// TIA Portal project "maupTIA_DEMO2023_V17" (V17) (continued)

       END_IF;
       #DrainingPhase.Cmd.StartMan := FALSE;
       #DrainingPhase.Cmd.PauseMan := FALSE;
       #DrainingPhase.Cmd.ResumeMan := FALSE;
       #DrainingPhase.Cmd.StopMan := FALSE;
   END_REGION

   REGION AutCtrl
       //if request to run in automatic mode -> set auto request to open of filling valve to 1 and close to 0, if not open 0 close 1
       // commands should be sets to false after their processing
       IF #DrainingPhase.State.AutCtrl THEN
           IF #DrainingPhase.Cmd.StartAut THEN
               #DrainingPhase.State.Running := TRUE;
               #DrainingPhase.State.Idle := FALSE;

               #DrainingPhase.Cmd.StartAut := FALSE;

               #DrainingValve.Cmd.AutCtrl := TRUE;




           END_IF;

           IF #DrainingPhase.Cmd.StopAut THEN
               #DrainingPhase.State.Running := FALSE;
               #DrainingPhase.State.Idle := TRUE;

               #DrainingPhase.Cmd.StopAut := FALSE;


           END_IF;

       END_IF;
   END_REGION

   REGION Done
       //every phase should have finish condition - draining phase - if water level is below requested level
       //after that done state should be setted to 1
       #DrainingPhase.Param.DrainLevel := 0.01;
       IF #DrainingPhase.WaterLevel <= #DrainingPhase.Param.DrainLevel THEN // kdyz je vypusteno, mozna je to zase ta promenna ktere preteka, nvm
           #DrainingPhase.Cmd.StopAut := TRUE;
           #DrainingPhase.Cmd.StopMan := TRUE;
           #DrainingPhase.State.Done := TRUE;
       END_IF;

       // command reset done resets done state and than resets command

       IF #DrainingPhase.Cmd.ResetDone THEN // AND DONE = TRUE? mozna zbytecne.
           #DrainingPhase.State.Done := FALSE;
           #DrainingPhase.Cmd.ResetDone := FALSE;
       END_IF;

   END_REGION

   REGION States 
       //Command valve in cases of states
       IF #DrainingPhase.State.Running THEN
           #DrainingValve.Cmd.Req2OpenAut := TRUE;
           #DrainingValve.Cmd.Req2CloseAut := FALSE;
          // #DrainingValve.Cmd.Req2CloseAut := FALSE;
       ELSE
           #DrainingValve.Cmd.Req2OpenAut := FALSE;
           #DrainingValve.Cmd.Req2CloseAut := TRUE;
           //#DrainingValve.Cmd.Req2CloseAut := FALSE;
       END_IF;
   END_REGION

   // delault state of phase - if not any state sets state to idle
   IF NOT #DrainingPhase.State.Idle AND NOT #DrainingPhase.State.Paused AND NOT #DrainingPhase.State.Running THEN
       #DrainingPhase.State.Idle := TRUE;
   END_IF;

   IF #DrainingPhase.State.Running THEN
       #DrainingPhase.State.StateInt := #Running;
   ELSIF #DrainingPhase.State.Paused THEN
       #DrainingPhase.State.StateInt := #Pause;
   ELSIF #DrainingPhase.State.Idle THEN
       #DrainingPhase.State.StateInt := #Idle;
   ELSIF #DrainingPhase.State.Done THEN
       #DrainingPhase.State.StateInt := #Idle;
   END_IF;
END_FUNCTION_BLOCK

FUNCTION_BLOCK "MixingFC"   // FB6, SCL
{ S7_Optimized_Access := 'TRUE' }
VERSION : 0.1
   VAR_IN_OUT
      MixingPhase : "PhaseMixing";
      MixerEng : "Engine";
   END_VAR
   VAR
      fElapsedTime : Int;
      fSecImp : R_TRIG;
   END_VAR
   VAR_TEMP
      tmp : Bool;
   END_VAR
   VAR CONSTANT
      Idle : Int := 0;
      Running : Int := 1;
      Pause : Int := 2;
   END_VAR
BEGIN
   REGION Aut/Man
       // switching state of engine - automatic or manual control (default state is manual)
       IF #MixingPhase.Cmd.AutCtrl THEN
           #MixingPhase.State.ManCtrl := FALSE;
           #MixingPhase.State.AutCtrl := TRUE;
           #MixingPhase.Cmd.AutCtrl := FALSE;
       END_IF;

       IF #MixingPhase.Cmd.ManCtrl THEN
           #MixingPhase.State.AutCtrl := FALSE;
           #MixingPhase.State.ManCtrl := TRUE;
           #MixingPhase.Cmd.ManCtrl := FALSE;
       END_IF;

       IF NOT #MixingPhase.State.AutCtrl AND NOT #MixingPhase.State.ManCtrl THEN
           #MixingPhase.State.ManCtrl := TRUE; // nebo dat Cmd.Manctrl do TRUE aby prosel IF nahore?
       END_IF;

   END_REGION

   REGION ManCtrl
       // processing manual actions - if command is processed, it is sets to FALSE even if can't be processed
       // Phase commands are start, stop, pause and resume 
       // Start - start mixing  
       // Stop - stop mixing
       // Pause - stop mixing 
       // Resume - start mixing
       // real states of phase are writed into states in phase structure

       IF #MixingPhase.State.ManCtrl THEN
           IF #MixingPhase.Cmd.StartMan THEN
               #MixingPhase.State.Paused := FALSE;
               #MixingPhase.State.Idle := FALSE;
               #MixingPhase.State.Running := TRUE;

               #MixerEng.Cmd.TurnOnMan := TRUE;
               //#MixerEng.Cmd.TurnOnMan := FALSE;

               #MixingPhase.Cmd.ResetDone := TRUE;
               //#MixingPhase.Cmd.ResetDone := FALSE;
           END_IF;

           IF #MixingPhase.State.Running THEN
               IF #MixingPhase.Cmd.PauseMan THEN
                   #MixingPhase.State.Running := FALSE;
                   #MixingPhase.State.Idle := FALSE;
                   #MixingPhase.State.Paused := TRUE;

                   #MixerEng.Cmd.TurnOffMan := TRUE;
                  // #MixerEng.Cmd.TurnOffMan := FALSE;

                   #MixingPhase.Cmd.ResetDone := TRUE;
                   //#MixingPhase.Cmd.ResetDone := FALSE;
               END_IF;
           END_IF;

           IF #MixingPhase.State.Paused THEN
               IF #MixingPhase.Cmd.ResumeMan THEN
                   #MixingPhase.State.Paused := FALSE;
                   #MixingPhase.State.Idle := FALSE;
                   #MixingPhase.State.Running := TRUE;

                   #MixerEng.Cmd.TurnOnMan := TRUE;
                   //#MixerEng.Cmd.TurnOnMan := FALSE;

                   #MixingPhase.Cmd.ResetDone := TRUE;
                   //#MixingPhase.Cmd.ResetDone := FALSE;
               END_IF;
           END_IF;


           IF #MixingPhase.State.Running OR #MixingPhase.State.Paused THEN
               IF #MixingPhase.Cmd.StopMan THEN
                   #MixingPhase.State.Running := FALSE;
                   #MixingPhase.State.Paused := FALSE;
                   #MixingPhase.State.Idle := TRUE;

                   #MixerEng.Cmd.TurnOffMan := TRUE;
                   //#MixerEng.Cmd.TurnOffMan := FALSE;

                   #MixingPhase.Cmd.ResetDone := TRUE;
                   //#MixingPhase.Cmd.ResetDone := FALSE;
               END_IF;
           END_IF;


       END_IF;
       #MixingPhase.Cmd.StartMan := FALSE;
       #MixingPhase.Cmd.PauseMan := FALSE;
       #MixingPhase.Cmd.ResumeMan := FALSE;
       #MixingPhase.Cmd.StopMan := FALSE;
   END_REGION

   REGION AutCtrl
       // if request to run in automatic mode -> set auto request to mixing to 1, if not request to mixing is 0
       // commands should be sets to false after their processing
       IF #MixingPhase.State.AutCtrl THEN
           IF #MixingPhase.Cmd.StartAut THEN
               #MixingPhase.State.Running := TRUE;
               #MixingPhase.State.Idle := FALSE;
               #MixingPhase.Cmd.StartAut := FALSE;
               #MixerEng.Cmd.AutCtrl := TRUE;
           END_IF;

           IF #MixingPhase.Cmd.StopAut THEN
               #MixingPhase.State.Running := FALSE;
               #MixingPhase.State.Idle := TRUE;
               #MixingPhase.Cmd.StopAut := FALSE;
           END_IF;

       END_IF;

   END_REGION


   REGION Done
       // every phase should have finish condition - mixing phase - if time of runnig is bigger or same as requested
       // after that done state should be setted to 1

       // command reset done resets done state and than resets command
       // calculation of elapsed time from engin state RT
       IF #MixingPhase.State.Running THEN
           "fSecImp"(CLK := "Clock_1Hz",
                     Q => #tmp);
           IF #tmp THEN
               #fElapsedTime := #fElapsedTime + 1;
           END_IF;

       END_IF;

       IF #MixingPhase.Param.TimeSec <= #fElapsedTime THEN // kdyz je domixovano, mozna je to zase ta promenna ktere preteka, nvm
           #MixingPhase.Cmd.StopAut := TRUE;
           #MixingPhase.Cmd.StopMan := TRUE;
           #MixingPhase.State.Done := TRUE;
       END_IF;


       // command reset done resets done state and than resets command
       IF #MixingPhase.Cmd.ResetDone THEN // AND DONE = TRUE? mozna zbytecne.
           // reset timer
           #MixingPhase.State.Done := FALSE;
           #fElapsedTime := 0;
           #MixingPhase.Cmd.ResetDone := FALSE;
       END_IF;


   END_REGION

   REGION States 
       //Command mixer in cases of states
    //??????????????
       IF #MixingPhase.State.Running THEN
           #MixerEng.Cmd.Req2RunAutCtrl := TRUE;
       ELSE
           #MixerEng.Cmd.Req2RunAutCtrl := FALSE;
       END_IF;
   END_REGION

   IF NOT #MixingPhase.State.Idle AND NOT #MixingPhase.State.Paused AND NOT #MixingPhase.State.Running THEN
       #MixingPhase.State.Idle := TRUE;
   END_IF;
   // delault state of phase - if not any state sets state to idle


   // delault state of phase - if not any state sets state to idle
   IF #MixingPhase.State.Running THEN
       #MixingPhase.State.StateInt := #Running;
   ELSIF #MixingPhase.State.Paused THEN
       #MixingPhase.State.StateInt := #Pause;
   ELSIF #MixingPhase.State.Idle THEN
       #MixingPhase.State.StateInt := #Idle;
   ELSIF #MixingPhase.State.Done THEN
       #MixingPhase.State.StateInt := #Idle;
   END_IF;
END_FUNCTION_BLOCK

FUNCTION_BLOCK "HeaterFC"   // FB7, SCL
{ S7_Optimized_Access := 'TRUE' }
VERSION : 0.1
   VAR_INPUT
      iWaterTemp : Real;
   END_VAR
   VAR_OUTPUT
      oHeaterEnable : Bool;
      oHeaterPower : Real;
   END_VAR
   VAR_IN_OUT
      iHeater_Struct : "Heater";
   END_VAR
   VAR
      fMode : Int;
   END_VAR
BEGIN
   #fMode := 3; // automatic mode of PID component
   "HeatingPID"(Setpoint := #iHeater_Struct.Param.HeatingSetPointAutomat,
                Input := #iWaterTemp,
                ManualEnable := #iHeater_Struct.State.ManCtrl,
                ManualValue := #iHeater_Struct.Param.HeatingPowerManual,
                OutputHeat => #iHeater_Struct.State.HeatingOut,
                Mode := #fMode);



   REGION Manual/Automat
       IF (NOT #iHeater_Struct.State.ManCtrl AND NOT #iHeater_Struct.State.AutCtrl) THEN
           #iHeater_Struct.State.ManCtrl := TRUE;
           #iHeater_Struct.State.AutCtrl := FALSE;
       ELSIF #iHeater_Struct.Cmd.ManCtrl THEN
           #iHeater_Struct.State.ManCtrl := TRUE;
           #iHeater_Struct.State.AutCtrl := FALSE;
           #iHeater_Struct.Cmd.ManCtrl := FALSE;
           #iHeater_Struct.Cmd.AutCtrl := FALSE;
       ELSIF #iHeater_Struct.Cmd.AutCtrl THEN
           #iHeater_Struct.State.ManCtrl := FALSE;
           #iHeater_Struct.State.AutCtrl := TRUE;
           #iHeater_Struct.Cmd.ManCtrl := FALSE;
           #iHeater_Struct.Cmd.AutCtrl := FALSE;
       END_IF;
   END_REGION

   REGION ManCtrl
       IF #iHeater_Struct.State.ManCtrl THEN
           IF #iHeater_Struct.Cmd.TurnOffMan THEN
               #iHeater_Struct.State.EnableOut := FALSE;
               #iHeater_Struct.Cmd.TurnOffMan := FALSE;
               #iHeater_Struct.Cmd.TurnOnMan := FALSE;
           ELSIF #iHeater_Struct.Cmd.TurnOnMan THEN
               #iHeater_Struct.State.EnableOut := TRUE;
               #iHeater_Struct.Cmd.TurnOffMan := FALSE;
               #iHeater_Struct.Cmd.TurnOnMan := FALSE;
           END_IF;
       END_IF;
   END_REGION

   REGION AutCtrl
       IF #iHeater_Struct.State.AutCtrl THEN
           #iHeater_Struct.State.EnableOut := #iHeater_Struct.Cmd.Req2RunAutCtrl;
       END_IF;
   END_REGION

   #oHeaterEnable := #iHeater_Struct.State.EnableOut;
   #oHeaterPower := #iHeater_Struct.State.HeatingOut;
END_FUNCTION_BLOCK

FUNCTION_BLOCK "Real2AnalogValue"   // FB8, SCL
{ S7_Optimized_Access := 'TRUE' }
VERSION : 0.1
   VAR_INPUT
      aiRealValue : Real;
      TransducerLoLevel : Int;
      TransducerHiLevel : Int;
      ScaledValLoLevel : Real;
      ScaledValHiLevel : Real;
   END_VAR
   VAR_OUTPUT
      aoRawAnalog : Int;
   END_VAR
BEGIN
   //#aoRawAnalog := (#TransducerHiLevel - #TransducerLoLevel) * REAL_TO_INT((#aiRealValue - #ScaledValLoLevel) / (#ScaledValHiLevel - #ScaledValLoLevel)) + #TransducerLoLevel;
   #aoRawAnalog := #TransducerLoLevel + REAL_TO_INT(#aiRealValue) * ((#TransducerHiLevel - #TransducerLoLevel) / REAL_TO_INT(#ScaledValHiLevel - #ScaledValLoLevel));
END_FUNCTION_BLOCK

FUNCTION_BLOCK "HeatingFC"   // FB9, SCL
{ S7_Optimized_Access := 'TRUE' }
VERSION : 0.1
   VAR_INPUT
      aiWaterTemp : Real;
   END_VAR
   VAR_IN_OUT
      HeatingPhase : "PhaseHeating";
      Heater : "Heater";
   END_VAR
   VAR
      fTime : Int;
      fSecImpEdge : R_TRIG;
   END_VAR
   VAR_TEMP
      tmp : Bool;
   END_VAR
   VAR CONSTANT
      Idle : Int := 0;
      Running : Int := 1;
      Pause : Int := 2;
   END_VAR
BEGIN
   REGION Aut/Man
       // switching state of engine - automatic or manual control (default state is manual)
       IF #HeatingPhase.Cmd.AutCtrl THEN
           #HeatingPhase.State.ManCtrl := FALSE;
           #HeatingPhase.State.AutCtrl := TRUE;
           #HeatingPhase.Cmd.AutCtrl := FALSE;
       END_IF;

       IF #HeatingPhase.Cmd.ManCtrl THEN
           #HeatingPhase.State.AutCtrl := FALSE;
           #HeatingPhase.State.ManCtrl := TRUE;
           #HeatingPhase.Cmd.ManCtrl := FALSE;
       END_IF;

       IF NOT #HeatingPhase.State.AutCtrl AND NOT #HeatingPhase.State.ManCtrl THEN
           #HeatingPhase.State.ManCtrl := TRUE; // nebo dat Cmd.Manctrl do TRUE aby prosel IF nahore?
           #HeatingPhase.State.AutCtrl := FALSE;
       END_IF;
   END_REGION

   REGION ManCtrl
       // processing manual actions - if command is processed, it is sets to FALSE even if can't be processed
       // real states of phase are writed into states in phase structure
       IF #HeatingPhase.State.ManCtrl THEN
           IF #HeatingPhase.Cmd.StartMan THEN
               #HeatingPhase.State.Paused := FALSE;
               #HeatingPhase.State.Idle := FALSE;
               #HeatingPhase.State.Running := TRUE;

               #Heater.Cmd.TurnOnMan := TRUE;
               #Heater.Cmd.TurnOnMan := FALSE;

               #HeatingPhase.Cmd.ResetDone := TRUE;
               #HeatingPhase.Cmd.ResetDone := FALSE;
           END_IF;

           IF #HeatingPhase.State.Running THEN
               IF #HeatingPhase.Cmd.PauseMan THEN
                   #HeatingPhase.State.Running := FALSE;
                   #HeatingPhase.State.Idle := FALSE;
                   #HeatingPhase.State.Paused := TRUE;

                   #Heater.Cmd.TurnOffMan := TRUE;
                   #Heater.Cmd.TurnOffMan := FALSE;

                   #HeatingPhase.Cmd.ResetDone := TRUE;
                   #HeatingPhase.Cmd.ResetDone := FALSE;
               END_IF;
           END_IF;

           IF #HeatingPhase.State.Paused THEN
               IF #HeatingPhase.Cmd.ResumeMan THEN
                   #HeatingPhase.State.Paused := FALSE;
                   #HeatingPhase.State.Idle := FALSE;
                   #HeatingPhase.State.Running := TRUE;

                   #Heater.Cmd.TurnOnMan := TRUE;
                   #Heater.Cmd.TurnOnMan := FALSE;

                   #HeatingPhase.Cmd.ResetDone := TRUE;
                   #HeatingPhase.Cmd.ResetDone := FALSE;
               END_IF;
           END_IF;


           IF #HeatingPhase.State.Running OR #HeatingPhase.State.Paused THEN
               IF #HeatingPhase.Cmd.StopMan THEN
                   #HeatingPhase.State.Running := FALSE;
                   #HeatingPhase.State.Paused := FALSE;
                   #HeatingPhase.State.Idle := TRUE;

                   #Heater.Cmd.TurnOffMan := TRUE;
                   #Heater.Cmd.TurnOffMan := FALSE;

                   #HeatingPhase.Cmd.ResetDone := TRUE;
                   #HeatingPhase.Cmd.ResetDone := FALSE;
               END_IF;
           END_IF;

       END_IF;
       #HeatingPhase.Cmd.StartMan := FALSE;
       #HeatingPhase.Cmd.PauseMan := FALSE;
       #HeatingPhase.Cmd.ResumeMan := FALSE;
       #HeatingPhase.Cmd.StopMan := FALSE; 
   END_REGION

   REGION AutCtrl
       // if request to run in automatic mode -> set auto request to heat to 1, if not request to heat 0
       // commands should be sets to false after their processing
       IF #HeatingPhase.State.AutCtrl THEN
           IF #HeatingPhase.Cmd.StartAut THEN
               #HeatingPhase.State.Running := TRUE;
               #HeatingPhase.State.Idle := FALSE;

               #HeatingPhase.Cmd.StartAut := FALSE;

               //#HeatingPhase.Cmd.AutCtrl := TRUE; // NEBO HO TAM DAT ROVNOU?
               //#HeatingPhase.Cmd.AutCtrl := FALSE;
           END_IF;

           IF #HeatingPhase.Cmd.StopAut THEN
               #HeatingPhase.State.Running := FALSE;
               #HeatingPhase.State.Idle := TRUE;
               #HeatingPhase.Cmd.StopAut := FALSE;
           END_IF;

       END_IF;
   END_REGION

   REGION Done
       //every phase should have finish condition - heating phase - if water temp is on requested value for 15 seconds with 1°C hysteresis
       //after that done state should be setted to 1
       ////AND #HeatingPhase.Param.ReqTemp <= #HeatingPhase.WaterTemp + 1 AND

       IF #HeatingPhase.State.Running THEN

           IF #HeatingPhase.Param.ReqTemp <= #HeatingPhase.WaterTemp THEN
               "fSecImp"(CLK := "Clock_1Hz",
                         Q => #tmp);
               IF #tmp THEN
                   #fTime := #fTime + 1;
               END_IF;

           END_IF;
           IF #fTime >= 10 THEN
               #HeatingPhase.State.Done := TRUE;
               #HeatingPhase.Cmd.StopAut := TRUE;
               #HeatingPhase.Cmd.StopMan := TRUE;
               #fTime := 0;
           END_IF;

       END_IF;

       (* IF #HeatingPhase.Param.ReqTemp = #aiWaterTemp THEN
           #HeatingPhase.Cmd.StopAut := TRUE;
           #HeatingPhase.Cmd.StopMan := TRUE;
           #HeatingPhase.State.Done := TRUE;
       END_IF; *)

       // command reset done resets done state and than resets command

       IF #HeatingPhase.Cmd.ResetDone THEN // AND DONE = TRUE? mozna zbytecne.
           #HeatingPhase.State.Done := FALSE;
           #HeatingPhase.Cmd.ResetDone := FALSE;
       END_IF;

   END_REGION

   REGION States 
       //Command valve in cases of states
       // Running - start heating  
       // Idle - stop heating
       // Pause - stop heating (alternative is hold actual temp)
       IF #HeatingPhase.State.Running THEN
           #Heater.Cmd.Req2RunAutCtrl := TRUE;
           #Heater.Param.HeatingSetPointAutomat := #HeatingPhase.Param.ReqTemp;
       END_IF;

       IF #HeatingPhase.State.Idle OR #HeatingPhase.State.Paused THEN
           #Heater.Cmd.Req2RunAutCtrl := FALSE;
       END_IF;


   END_REGION

   IF NOT #HeatingPhase.State.Idle AND NOT #HeatingPhase.State.Paused AND NOT #HeatingPhase.State.Running THEN
       #HeatingPhase.State.Idle := TRUE;
   END_IF;
   // delault state of phase - if not any state sets state to idle

   IF #HeatingPhase.State.Running THEN
       #HeatingPhase.State.StateInt := #Running;
   ELSIF #HeatingPhase.State.Paused THEN
       #HeatingPhase.State.StateInt := #Pause;
   ELSIF #HeatingPhase.State.Idle THEN
       #HeatingPhase.State.StateInt := #Idle;
   ELSIF #HeatingPhase.State.Done THEN
       #HeatingPhase.State.StateInt := #Idle;
   END_IF;
END_FUNCTION_BLOCK

FUNCTION "AnalogScalingFC" : Void   // FC1, SCL
{ S7_Optimized_Access := 'TRUE' }
VERSION : 0.1
   VAR_INPUT
      aiRAWanalog : Int;
      TransducerLoLevel : Int;
      TransducerHiLevel : Int;
      ScaledValLoLevel : Real;
      ScaledValHiLevel : Real;
   END_VAR
   VAR_OUTPUT
      aoScaledValue : Real;
   END_VAR
   VAR_IN_OUT
      PrevVal : Real;
   END_VAR
   VAR_TEMP
      NormValue : Real;
      LastVal : Real;
   END_VAR
BEGIN
   //#aoScaledValue := (#ScaledValHiLevel - #ScaledValLoLevel) * ((INT_TO_REAL(#aiRAWanalog - #TransducerLoLevel)) / (INT_TO_REAL(#TransducerHiLevel - #TransducerLoLevel))) + #ScaledValLoLevel;

   #NormValue := NORM_X(MIN := #TransducerLoLevel, VALUE := #aiRAWanalog, MAX := #TransducerHiLevel);

   #aoScaledValue := SCALE_X(MIN := #ScaledValLoLevel, VALUE := #NormValue, MAX := #ScaledValHiLevel);

   IF #LastVal = #LastVal THEN
       #LastVal := #LastVal;
   ELSE
       #LastVal := 0; 
   END_IF;


   IF (#aoScaledValue-#PrevVal) < (0.95*#ScaledValHiLevel)THEN
       #aoScaledValue := #aoScaledValue;
       // ulozeni nove hodnoty do minule pro dalsi porovnani
       #PrevVal := #aoScaledValue;

   END_IF;

   IF (#aoScaledValue-#PrevVal) > (0.95*#ScaledValHiLevel) THEN
       #aoScaledValue := #PrevVal;
   END_IF;
END_FUNCTION

(* ===== HMI "HMI_RT_1" =====
system functions are stored by id; their names below are inferred from use
connection "HMI_Connection_2": ETHERNET, S7_1500_OMS

HMI tags "Default tag table"
   "Tag_ScreenNumber" : UInt, internal
   "Data_Tank1_ValveFill_State_AutCtrl" : Bool = PLC Data.Tank1.ValveFill.State.AutCtrl, 100 ms
   "Data_Tank1_ValveFill_State_ManCtrl" : Bool = PLC Data.Tank1.ValveFill.State.ManCtrl, 100 ms
   "Data_Tank1_ValveFill_State_Open" : Bool = PLC Data.Tank1.ValveFill.State.Open, 100 ms
   "Data_Tank1_ValveFill_State_Closed" : Bool = PLC Data.Tank1.ValveFill.State.Closed, 100 ms
   "Data_Tank1_Mixer_State_AutCtrl" : Bool = PLC Data.Tank1.Mixer.State.AutCtrl, 100 ms
   "Data_Tank1_Mixer_State_ManCtrl" : Bool = PLC Data.Tank1.Mixer.State.ManCtrl, 100 ms
   "Data_Tank1_Mixer_State_Run" : Bool = PLC Data.Tank1.Mixer.State.Run, 100 ms
   "Data_Tank1_ValveDrain_State_AutCtrl" : Bool = PLC Data.Tank1.ValveDrain.State.AutCtrl, 100 ms
   "Data_Tank1_ValveDrain_State_ManCtrl" : Bool = PLC Data.Tank1.ValveDrain.State.ManCtrl, 100 ms
   "Data_Tank1_ValveDrain_State_Open" : Bool = PLC Data.Tank1.ValveDrain.State.Open, 100 ms
   "Data_Tank1_ValveDrain_State_Closed" : Bool = PLC Data.Tank1.ValveDrain.State.Closed, 100 ms
   "Data_Tank1_ValveFill_Cmd_AutCtrl" : Bool = PLC Data.Tank1.ValveFill.Cmd.AutCtrl, 100 ms
   "Data_Tank1_ValveFill_Cmd_ManCtrl" : Bool = PLC Data.Tank1.ValveFill.Cmd.ManCtrl, 100 ms
   "Data_Tank1_ValveFill_Cmd_OpenMan" : Bool = PLC Data.Tank1.ValveFill.Cmd.OpenMan, 100 ms
   "Data_Tank1_ValveFill_Cmd_CloseMan" : Bool = PLC Data.Tank1.ValveFill.Cmd.CloseMan, 100 ms
   "Data_Tank1_Mixer_Cmd_AutCtrl" : Bool = PLC Data.Tank1.Mixer.Cmd.AutCtrl, 100 ms
   "Data_Tank1_Mixer_Cmd_ManCtrl" : Bool = PLC Data.Tank1.Mixer.Cmd.ManCtrl, 100 ms
   "Data_Tank1_Mixer_Cmd_TurnOnMan" : Bool = PLC Data.Tank1.Mixer.Cmd.TurnOnMan, 100 ms
   "Data_Tank1_Mixer_Cmd_TurnOffMan" : Bool = PLC Data.Tank1.Mixer.Cmd.TurnOffMan, 100 ms
   "Data_Tank1_ValveDrain_Cmd_AutCtrl" : Bool = PLC Data.Tank1.ValveDrain.Cmd.AutCtrl, 100 ms
   "Data_Tank1_ValveDrain_Cmd_OpenMan" : Bool = PLC Data.Tank1.ValveDrain.Cmd.OpenMan, 100 ms
   "Data_Tank1_ValveDrain_Cmd_CloseMan" : Bool = PLC Data.Tank1.ValveDrain.Cmd.CloseMan, 100 ms
   "Data_Tank1_WaterLevel_AIScaled" : Real = PLC Data.Tank1.WaterLevel.AIScaled, 100 ms
   "Data_Tank1_WaterTemp_AIScaled" : Real = PLC Data.Tank1.WaterTemp.AIScaled, 100 ms
   "HeatingPID_ManualEnable" : Bool = PLC HeatingPID.ManualEnable, 100 ms
   "Data_Tank1_Heating_Param_ReqTemp" : Real = PLC Data.Tank1.Heating.Param.ReqTemp, 100 ms
   "Data_Tank1_Filling_State_Stateint" : Int = PLC Data.Tank1.Filling.State.Stateint, 100 ms
   "Data_Tank1_Draining_State_StateInt" : Int = PLC Data.Tank1.Draining.State.StateInt, 100 ms
   "Data_Tank1_Mixing_State_StateInt" : Int = PLC Data.Tank1.Mixing.State.StateInt, 100 ms
   "Data_Tank1_Heating_State_StateInt" : Int = PLC Data.Tank1.Heating.State.StateInt, 100 ms
   "Data_Tank1_Filling_State_AutCtrl" : Bool = PLC Data.Tank1.Filling.State.AutCtrl, 100 ms
   "Data_Tank1_Filling_State_ManCtrl" : Bool = PLC Data.Tank1.Filling.State.ManCtrl, 100 ms
   "Data_Tank1_Filling_State_Done" : Bool = PLC Data.Tank1.Filling.State.Done, 100 ms
   "Data_Tank1_Filling_Cmd_AutCtrl" : Bool = PLC Data.Tank1.Filling.Cmd.AutCtrl, 100 ms
   "Data_Tank1_Filling_Cmd_ManCtrl" : Bool = PLC Data.Tank1.Filling.Cmd.ManCtrl, 100 ms
   "Data_Tank1_Filling_Cmd_ResetDone" : Bool = PLC Data.Tank1.Filling.Cmd.ResetDone, 100 ms
   "Data_Tank1_Filling_Cmd_StartMan" : Bool = PLC Data.Tank1.Filling.Cmd.StartMan, 100 ms
   "Data_Tank1_Filling_Cmd_StopMan" : Bool = PLC Data.Tank1.Filling.Cmd.StopMan, 100 ms
   "Data_Tank1_Filling_Cmd_PauseMan" : Bool = PLC Data.Tank1.Filling.Cmd.PauseMan, 100 ms
   "Data_Tank1_Filling_Cmd_ResumeMan" : Bool = PLC Data.Tank1.Filling.Cmd.ResumeMan, 100 ms
   "Data_Tank1_Mixing_State_AutCtrl" : Bool = PLC Data.Tank1.Mixing.State.AutCtrl, 100 ms
   "Data_Tank1_Mixing_State_ManCtrl" : Bool = PLC Data.Tank1.Mixing.State.ManCtrl, 100 ms
   "Data_Tank1_Mixing_State_Done" : Bool = PLC Data.Tank1.Mixing.State.Done, 100 ms
   "Data_Tank1_Mixing_Cmd_AutCtrl" : Bool = PLC Data.Tank1.Mixing.Cmd.AutCtrl, 100 ms
   "Data_Tank1_Mixing_Cmd_ManCtrl" : Bool = PLC Data.Tank1.Mixing.Cmd.ManCtrl, 100 ms
   "Data_Tank1_Mixing_Cmd_ResetDone" : Bool = PLC Data.Tank1.Mixing.Cmd.ResetDone, 100 ms
   "Data_Tank1_Mixing_Cmd_StartMan" : Bool = PLC Data.Tank1.Mixing.Cmd.StartMan, 100 ms
   "Data_Tank1_Mixing_Cmd_StopMan" : Bool = PLC Data.Tank1.Mixing.Cmd.StopMan, 100 ms
   "Data_Tank1_Mixing_Cmd_PauseMan" : Bool = PLC Data.Tank1.Mixing.Cmd.PauseMan, 100 ms
   "Data_Tank1_Mixing_Cmd_ResumeMan" : Bool = PLC Data.Tank1.Mixing.Cmd.ResumeMan, 100 ms
   "Data_Tank1_Draining_State_AutCtrl" : Bool = PLC Data.Tank1.Draining.State.AutCtrl, 100 ms
   "Data_Tank1_Draining_State_ManCtrl" : Bool = PLC Data.Tank1.Draining.State.ManCtrl, 100 ms
   "Data_Tank1_Draining_State_Done" : Bool = PLC Data.Tank1.Draining.State.Done, 100 ms
   "Data_Tank1_Draining_Cmd_AutCtrl" : Bool = PLC Data.Tank1.Draining.Cmd.AutCtrl, 100 ms
   "Data_Tank1_Draining_Cmd_ManCtrl" : Bool = PLC Data.Tank1.Draining.Cmd.ManCtrl, 100 ms
   "Data_Tank1_Draining_Cmd_ResetDone" : Bool = PLC Data.Tank1.Draining.Cmd.ResetDone, 100 ms
   "Data_Tank1_Draining_Cmd_StartMan" : Bool = PLC Data.Tank1.Draining.Cmd.StartMan, 100 ms
   "Data_Tank1_Draining_Cmd_StopMan" : Bool = PLC Data.Tank1.Draining.Cmd.StopMan, 100 ms
   "Data_Tank1_Draining_Cmd_PauseMan" : Bool = PLC Data.Tank1.Draining.Cmd.PauseMan, 100 ms
   "Data_Tank1_Draining_Cmd_ResumeMan" : Bool = PLC Data.Tank1.Draining.Cmd.ResumeMan, 100 ms
   "Data_Tank1_Heating_State_AutCtrl" : Bool = PLC Data.Tank1.Heating.State.AutCtrl, 100 ms
   "Data_Tank1_Heating_State_ManCtrl" : Bool = PLC Data.Tank1.Heating.State.ManCtrl, 100 ms
   "Data_Tank1_Heating_State_Done" : Bool = PLC Data.Tank1.Heating.State.Done, 100 ms
   "Data_Tank1_Heating_Cmd_AutCtrl" : Bool = PLC Data.Tank1.Heating.Cmd.AutCtrl, 100 ms
   "Data_Tank1_Heating_Cmd_ManCtrl" : Bool = PLC Data.Tank1.Heating.Cmd.ManCtrl, 100 ms
   "Data_Tank1_Heating_Cmd_ResetDone" : Bool = PLC Data.Tank1.Heating.Cmd.ResetDone, 100 ms
   "Data_Tank1_Heating_Cmd_StartMan" : Bool = PLC Data.Tank1.Heating.Cmd.StartMan, 100 ms
   "Data_Tank1_Heating_Cmd_StopMan" : Bool = PLC Data.Tank1.Heating.Cmd.StopMan, 100 ms
   "Data_Tank1_Heating_Cmd_PauseMan" : Bool = PLC Data.Tank1.Heating.Cmd.PauseMan, 100 ms
   "Data_Tank1_Heating_Cmd_ResumeMan" : Bool = PLC Data.Tank1.Heating.Cmd.ResumeMan, 100 ms
   "Data_Tank1_Filling_Param_FillLevel" : Real = PLC Data.Tank1.Filling.Param.FillLevel, 100 ms
   "Data_Tank1_Draining_Param_DrainLevel" : Real = PLC Data.Tank1.Draining.Param.DrainLevel, 100 ms
   "Data_Tank1_Mixing_Param_TimeSec" : Int = PLC Data.Tank1.Mixing.Param.TimeSec, 100 ms
   "Data_Tank1_Mixer_State_StateInt" : Int = PLC Data.Tank1.Mixer.State.StateInt, 100 ms
   "Data_Tank1_ValveFill_State_StColor" : Int = PLC Data.Tank1.ValveFill.State.StColor, 100 ms
   "Data_Tank1_ValveDrain_State_StColor" : Int = PLC Data.Tank1.ValveDrain.State.StColor, 100 ms
   "Data_Tank1_ValveDrain_Cmd_ManCtrl" : Bool = PLC Data.Tank1.ValveDrain.Cmd.ManCtrl, 100 ms
   "Data_Tank1_Heater_Cmd_AutCtrl" : Bool = PLC Data.Tank1.Heater.Cmd.AutCtrl, 100 ms
   "Data_Tank1_Heater_Cmd_ManCtrl" : Bool = PLC Data.Tank1.Heater.Cmd.ManCtrl, 100 ms
   "Data_Tank1_Heater_Cmd_TurnOnMan" : Bool = PLC Data.Tank1.Heater.Cmd.TurnOnMan, 100 ms
   "Data_Tank1_Heater_Cmd_TurnOffMan" : Bool = PLC Data.Tank1.Heater.Cmd.TurnOffMan, 100 ms
   "Data_Tank1_Heater_Param_HeatingPowerManual" : Real = PLC Data.Tank1.Heater.Param.HeatingPowerManual, 100 ms
   "Data_Tank1_Heater_State_AutCtrl" : Bool = PLC Data.Tank1.Heater.State.AutCtrl, 100 ms
   "Data_Tank1_Heater_State_ManCtrl" : Bool = PLC Data.Tank1.Heater.State.ManCtrl, 100 ms
   "Data_Tank1_Mixing_Cmd_Auto_Start" : Bool = PLC Data.Tank1.Mixing.Cmd.StartAut AT %DB1.DBX0.0, 1 s
   "Data_Tank1_Mixing_Cmd_Auto_Stop" : Bool = PLC Data.Tank1.Mixing.Cmd.StopAut AT %DB1.DBX0.0, 1 s

text list "Phases": 0 'Idle'; 1 'Running'; 2 'Pause'

text list "Process": 0 'Running'; 1 'Idle'; 2 'Stopping'

screen "MainScr" 800x480
   SymbolLibrary "Symbol library_1" at 202,63 size 120x212
   SymbolLibrary "Symbol library_2" at 148,84 size 58x23
   SymbolLibrary "Symbol library_3" at 320,241 size 20x23
   Bar "Bar_1" at 204,63 size 117x211; MinimumValue 0; MaximumValue 2
      ProcessValue <- "Data_Tank1_WaterLevel_AIScaled"
   SymbolLibrary "Symbol library_4" at 55,31 size 94x80
      Appearance <- "Data_Tank1_ValveFill_State_StColor"
   IOField "I/O field_1" at 215,109 size 96x32; FormatPattern s9.99; Unit  m
      ProcessValue <- "Data_Tank1_WaterLevel_AIScaled"
   IOField "I/O field_2" at 216,143 size 96x32; FormatPattern 999.9; Unit  °C
      ProcessValue <- "Data_Tank1_WaterTemp_AIScaled"
   SymbolLibrary "Symbol library_6" at 226,190 size 71x61
      Appearance <- "Data_Tank1_Mixer_State_StateInt"
   Button "Button_1" at 17,393 size 77x32; TextOff 'Aut'
      on Click: SetBit("Data_Tank1_ValveFill_Cmd_AutCtrl")
   TextField "Text field_1" at 55,283 size 83x23; Text 'ValveFill'
   TextField "Text field_2" at 15,308 size 83x23; Text 'Automat'
   TextField "Text field_3" at 15,326 size 70x23; Text 'Manual'
   TextField "Text field_4" at 15,348 size 51x23; Text 'Open'
   TextField "Text field_5" at 15,366 size 65x23; Text 'Closed'
   Button "Button_2" at 96,393 size 77x32; TextOff 'Man'
      on Click: SetBit("Data_Tank1_ValveFill_Cmd_ManCtrl")
   Button "Button_3" at 17,427 size 77x32; TextOff 'Open'
      on Click: SetBit("Data_Tank1_ValveFill_Cmd_OpenMan")
   Button "Button_4" at 96,427 size 77x32; TextOff 'Close'
      on Click: SetBit("Data_Tank1_ValveFill_Cmd_CloseMan")
   Circle "Circle_1" at 132,309 size 20x20
      Appearance <- "Data_Tank1_ValveFill_State_AutCtrl"
   Circle "Circle_2" at 132,329 size 20x20
      Appearance <- "Data_Tank1_ValveFill_State_ManCtrl"
   Circle "Circle_3" at 132,349 size 20x20
      Appearance <- "Data_Tank1_ValveFill_State_Open"
   Circle "Circle_4" at 132,369 size 20x20
      Appearance <- "Data_Tank1_ValveFill_State_Closed"
   TextField "Text field_6" at 450,99 size 104x23; Text 'ValveDrain'
   TextField "Text field_7" at 417,124 size 83x23; Text 'Automat'
   TextField "Text field_8" at 417,142 size 70x23; Text 'Manual'
   TextField "Text field_9" at 417,164 size 51x23; Text 'Open'
   TextField "Text field_10" at 417,182 size 65x23; Text 'Closed'
   TextField "Text field_11" at 234,284 size 56x23; Text 'Mixer'
   TextField "Text field_12" at 185,309 size 83x23; Text 'Automat'
   TextField "Text field_13" at 185,327 size 70x23; Text 'Manual'
   TextField "Text field_14" at 185,350 size 79x23; Text 'Running'
   Circle "Circle_9" at 302,310 size 20x20
      Appearance <- "Data_Tank1_Mixer_State_AutCtrl"
   Circle "Circle_10" at 302,330 size 20x20
      Appearance <- "Data_Tank1_Mixer_State_ManCtrl"
   Circle "Circle_12" at 302,354 size 20x20
      Appearance <- "Data_Tank1_Mixer_State_Run"
   TextField "Text field_16" at 662,99 size 77x27; Text 'Phases'
   Button "Button_15" at 617,148 size 171x29; TextOff 'Menu filling'
      on Click: ActivateScreen("Filling", 0)
   TextField "Text field_17" at 668,124 size 61x23; Text 'Filling'
   SymbolicIOField "Symbolic I/O field_2" at 617,179 size 171x32; TextOn '1'; TextOff '0'; TextList "Phases"
      ProcessValue <- "Data_Tank1_Filling_State_Stateint"
   Button "Button_16" at 617,236 size 171x29; TextOff 'Menu draining'
      on Click: ActivateScreen("Draining", 0)
   TextField "Text field_18" at 660,213 size 82x23; Text 'Draining'
   SymbolicIOField "Symbolic I/O field_3" at 617,267 size 171x32; TextOn '1'; TextOff '0'; TextList "Phases"
      ProcessValue <- "Data_Tank1_Draining_State_StateInt"
   Button "Button_17" at 617,324 size 171x29; TextOff 'Menu mixing'
      on Click: ActivateScreen("Mixing", 0)
   TextField "Text field_19" at 669,301 size 65x23; Text 'Mixing'
   SymbolicIOField "Symbolic I/O field_4" at 617,355 size 171x32; TextOn '1'; TextOff '0'; TextList "Phases"
      ProcessValue <- "Data_Tank1_Mixing_State_StateInt"
   Button "Button_18" at 617,412 size 171x29; TextOff 'Menu heating'
      on Click: ActivateScreen("Heating", 0)
   TextField "Text field_20" at 665,390 size 76x23; Text 'Heating'
   SymbolicIOField "Symbolic I/O field_5" at 617,443 size 171x32; TextOn '1'; TextOff '0'; TextList "Phases"
      ProcessValue <- "Data_Tank1_Heating_State_StateInt"
   TextField "Text field_21" at 427,285 size 156x23; Text 'Heating element'
   TextField "Text field_22" at 418,310 size 83x23; Text 'Automat'
   TextField "Text field_23" at 418,328 size 70x23; Text 'Manual'
   TextField "Text field_24" at 422,350 size 157x23; Text 'Manual heat pwr'
   IOField "I/O field_3" at 447,371 size 96x32; FormatPattern s999.99; Unit  %
      Appearance <- "Data_Tank1_Heater_Param_HeatingPowerManual"
      ProcessValue <- "Data_Tank1_Heater_Param_HeatingPowerManual"
   Button "Button_19" at 335,12 size 130x66; TextOff 'Parameters tank 1'
      on Click: ActivateScreen("Parameters", 0)
   Button "Button_5" at 416,208 size 77x32; TextOff 'Aut'
      on Click: SetBit("Data_Tank1_ValveDrain_Cmd_AutCtrl")
   Button "Button_6" at 503,207 size 77x32; TextOff 'Man'
      on Click: SetBit("Data_Tank1_ValveDrain_Cmd_ManCtrl")
   Button "Button_7" at 416,242 size 77x32; TextOff 'Open'
      on Click: SetBit("Data_Tank1_ValveDrain_Cmd_OpenMan")
   Button "Button_8" at 503,242 size 77x32; TextOff 'Close'
      on Click: SetBit("Data_Tank1_ValveDrain_Cmd_CloseMan")
   Circle "Circle_5" at 536,128 size 20x20
      Appearance <- "Data_Tank1_ValveDrain_State_AutCtrl"
   Circle "Circle_6" at 536,147 size 20x20
      Appearance <- "Data_Tank1_ValveDrain_State_ManCtrl"
   Circle "Circle_7" at 536,166 size 20x20
      Appearance <- "Data_Tank1_ValveDrain_State_Open"
   Circle "Circle_8" at 536,186 size 20x20
      Appearance <- "Data_Tank1_ValveDrain_State_Closed"
   Button "Button_9" at 187,380 size 77x32; TextOff 'Aut'
      on Click: SetBit("Data_Tank1_Mixer_Cmd_AutCtrl")
   Button "Button_10" at 187,412 size 77x32; TextOff 'On'
      on Click: SetBit("Data_Tank1_Mixer_Cmd_TurnOnMan")
   Button "Button_11" at 268,381 size 77x32; TextOff 'Man'
      on Click: SetBit("Data_Tank1_Mixer_Cmd_ManCtrl")
   Button "Button_12" at 268,412 size 77x32; TextOff 'Off'
      on Click: SetBit("Data_Tank1_Mixer_Cmd_TurnOffMan")
   Circle "Circle_11" at 538,313 size 20x20
      Appearance <- "Data_Tank1_Heater_State_AutCtrl"
   Circle "Circle_13" at 538,332 size 20x20
      Appearance <- "Data_Tank1_Heater_State_ManCtrl"
   Button "Button_13" at 418,402 size 77x32; TextOff 'Aut'
      on Click: SetBit("Data_Tank1_Heater_Cmd_AutCtrl")
   Button "Button_14" at 501,402 size 77x32; TextOff 'Man'
      on Click: SetBit("Data_Tank1_Heater_Cmd_ManCtrl")
   Button "Button_20" at 418,433 size 77x32; TextOff 'On'
      on Click: SetBit("Data_Tank1_Heater_Cmd_TurnOnMan")
   Button "Button_21" at 501,434 size 77x32; TextOff 'Off'
      on Click: SetBit("Data_Tank1_Heater_Cmd_TurnOffMan")
   SymbolLibrary "Symbol library_5" at 311,188 size 94x80
      Appearance <- "Data_Tank1_ValveDrain_State_StColor"

screen "Heating" 800x480
   TextField "Text field_26" at 278,299 size 205x23; Text 'Heating phase control'
   TextField "Text field_27" at 182,333 size 83x23; Text 'Automat'
   TextField "Text field_28" at 182,351 size 70x23; Text 'Manual'
   TextField "Text field_29" at 343,342 size 51x23; Text 'Done'
   GraphicView "Graphic view_1" at 525,294 size 75x74; Picture "exit-png-cancel-cross-exit-remove-icon-512"
   Button "Button_26" at 520,296 size 76x81; TextOff 'Text'
      on Click: ActivateScreen("MainScr", 0)
   Button "Button_5" at 185,385 size 77x32; TextOff 'Aut'
      on Click: SetBit("Data_Tank1_Heating_Cmd_AutCtrl")
   Button "Button_6" at 185,422 size 77x32; TextOff 'Start'
      on Click: SetBit("Data_Tank1_Heating_Cmd_StartMan")
   Button "Button_7" at 262,385 size 77x32; TextOff 'Man'
      on Click: SetBit("Data_Tank1_Heating_Cmd_ManCtrl")
   Button "Button_13" at 262,422 size 77x32; TextOff 'Stop'
      on Click: SetBit("Data_Tank1_Heating_Cmd_StopMan")
   Button "Button_8" at 340,385 size 158x32; TextOff 'Reset Done'
      on Click: SetBit("Data_Tank1_Heating_Cmd_ResetDone")
   Button "Button_14" at 345,422 size 77x32; TextOff 'Pause'
      on Click: SetBit("Data_Tank1_Heating_Cmd_PauseMan")
   Button "Button_19" at 422,422 size 77x32; TextOff 'Rsume'
      on Click: SetBit("Data_Tank1_Heating_Cmd_ResumeMan")
   Circle "Circle_5" at 433,336 size 35x35
      Appearance <- "Data_Tank1_Heating_State_Done"
   Circle "Circle_6" at 291,336 size 20x20
      Appearance <- "Data_Tank1_Heating_State_AutCtrl"
   Circle "Circle_7" at 292,353 size 20x20
      Appearance <- "Data_Tank1_Heating_State_ManCtrl"
   SymbolLibrary "Symbol library_1" at 202,63 size 120x212
   SymbolLibrary "Symbol library_2" at 148,84 size 58x23
   SymbolLibrary "Symbol library_3" at 320,241 size 20x23
   Bar "Bar_1" at 204,63 size 117x211; MinimumValue 0; MaximumValue 2
      ProcessValue <- "Data_Tank1_WaterLevel_AIScaled"
   SymbolLibrary "Symbol library_4" at 55,31 size 94x80
      Appearance <- "Data_Tank1_ValveFill_State_StColor"
   IOField "I/O field_1" at 215,109 size 96x32; FormatPattern s9.99; Unit  m
      ProcessValue <- "Data_Tank1_WaterLevel_AIScaled"
   IOField "I/O field_2" at 216,143 size 96x32; FormatPattern 999.9; Unit  °C
      ProcessValue <- "Data_Tank1_WaterTemp_AIScaled"
   SymbolLibrary "Symbol library_6" at 226,190 size 71x61
      Appearance <- "Data_Tank1_Mixer_State_StateInt"
   Button "Button_1" at 7,233 size 77x32; TextOff 'Aut'
      on Click: SetBit("Data_Tank1_ValveFill_Cmd_AutCtrl")
   TextField "Text field_1" at 45,123 size 83x23; Text 'ValveFill'
   TextField "Text field_2" at 5,148 size 83x23; Text 'Automat'
   TextField "Text field_3" at 5,166 size 70x23; Text 'Manual'
   TextField "Text field_4" at 5,188 size 51x23; Text 'Open'
   TextField "Text field_5" at 5,206 size 65x23; Text 'Closed'
   Button "Button_2" at 86,233 size 77x32; TextOff 'Man'
      on Click: SetBit("Data_Tank1_ValveFill_Cmd_ManCtrl")
   Button "Button_3" at 7,267 size 77x32; TextOff 'Open'
      on Click: SetBit("Data_Tank1_ValveFill_Cmd_OpenMan")
   Button "Button_4" at 86,267 size 77x32; TextOff 'Close'
      on Click: SetBit("Data_Tank1_ValveFill_Cmd_CloseMan")
   TextField "Text field_6" at 450,99 size 104x23; Text 'ValveDrain'
   TextField "Text field_7" at 417,124 size 83x23; Text 'Automat'
   TextField "Text field_8" at 417,142 size 70x23; Text 'Manual'
   TextField "Text field_9" at 417,164 size 51x23; Text 'Open'
   TextField "Text field_10" at 417,182 size 65x23; Text 'Closed'
   Button "Button_9" at 187,378 size 77x32; TextOff 'Aut'
      on Click: SetBit("Data_Tank1_Mixer_Cmd_AutCtrl")
   TextField "Text field_11" at 234,284 size 56x23; Text 'Mixer'
   TextField "Text field_12" at 185,309 size 83x23; Text 'Automat'
   TextField "Text field_13" at 185,327 size 70x23; Text 'Manual'
   TextField "Text field_14" at 185,350 size 79x23; Text 'Running'
   Button "Button_10" at 266,378 size 77x32; TextOff 'Man'
      on Click: SetBit("Data_Tank1_Mixer_Cmd_ManCtrl")
   Button "Button_11" at 187,411 size 77x32; TextOff 'Start'
      on Click: SetBit("Data_Tank1_Mixer_Cmd_TurnOnMan")
   Button "Button_12" at 266,411 size 77x32; TextOff 'Stop'
      on Click: SetBit("Data_Tank1_Mixer_Cmd_TurnOffMan")
   TextField "Text field_16" at 662,99 size 77x27; Text 'Phases'
   Button "Button_15" at 617,148 size 171x29; TextOff 'Menu filling'
      on Click: ActivateScreen("Filling", 0)
   TextField "Text field_17" at 668,124 size 61x23; Text 'Filling'
   SymbolicIOField "Symbolic I/O field_2" at 617,179 size 171x32; TextOn '1'; TextOff '0'; TextList "Phases"
      ProcessValue <- "Data_Tank1_Filling_State_Stateint"
   Button "Button_16" at 617,236 size 171x29; TextOff 'Menu draining'
      on Click: ActivateScreen("Draining", 0)
   TextField "Text field_18" at 660,213 size 82x23; Text 'Draining'
   SymbolicIOField "Symbolic I/O field_3" at 617,267 size 171x32; TextOn '1'; TextOff '0'; TextList "Phases"
      ProcessValue <- "Data_Tank1_Draining_State_StateInt"
   Button "Button_17" at 617,324 size 171x29; TextOff 'Menu mixing'
      on Click: ActivateScreen("Mixing", 0)
   TextField "Text field_19" at 669,301 size 65x23; Text 'Mixing'
   SymbolicIOField "Symbolic I/O field_4" at 617,355 size 171x32; TextOn '1'; TextOff '0'; TextList "Phases"
      ProcessValue <- "Data_Tank1_Mixing_State_StateInt"
   Button "Button_18" at 617,412 size 171x29; TextOff 'Menu heating'
      on Click: ActivateScreen("Heating", 0)
   TextField "Text field_20" at 665,390 size 76x23; Text 'Heating'
   SymbolicIOField "Symbolic I/O field_5" at 617,443 size 171x32; TextOn '1'; TextOff '0'; TextList "Phases"
      ProcessValue <- "Data_Tank1_Heating_State_StateInt"
   TextField "Text field_21" at 427,291 size 156x23; Text 'Heating element'
   TextField "Text field_22" at 418,316 size 83x23; Text 'Automat'
   TextField "Text field_23" at 418,334 size 70x23; Text 'Manual'
   TextField "Text field_24" at 422,356 size 157x23; Text 'Manual heat pwr'
   IOField "I/O field_3" at 447,377 size 96x32; FormatPattern 999.9; Unit  %
      ProcessValue <- "Data_Tank1_Heater_Param_HeatingPowerManual"
   TextField "Text field_25" at 422,408 size 160x23; Text 'Req temperature'
   IOField "I/O field_4" at 447,429 size 96x32; FormatPattern 999.9; Unit  °C
      ProcessValue <- "Data_Tank1_Heating_Param_ReqTemp"
   Button "Button_27" at 335,12 size 130x66; TextOff 'Parameters tank 1'
      on Click: ActivateScreen("Parameters", 0)
   Circle "Circle_1" at 122,149 size 20x20
      Appearance <- "Data_Tank1_ValveFill_State_AutCtrl"
   Circle "Circle_2" at 122,169 size 20x20
      Appearance <- "Data_Tank1_ValveFill_State_ManCtrl"
   Circle "Circle_3" at 122,189 size 20x20
      Appearance <- "Data_Tank1_ValveFill_State_Open"
   Circle "Circle_4" at 122,209 size 20x20
      Appearance <- "Data_Tank1_ValveFill_State_Closed"
   Circle "Circle_9" at 302,310 size 20x20
      Appearance <- "Data_Tank1_Mixer_State_AutCtrl"
   Circle "Circle_10" at 302,330 size 20x20
      Appearance <- "Data_Tank1_Mixer_State_ManCtrl"
   Circle "Circle_12" at 302,354 size 20x20
      Appearance <- "Data_Tank1_Mixer_State_Run"
   Circle "Circle_11" at 535,317 size 20x20
      Appearance <- "Data_Tank1_Heating_Cmd_AutCtrl"
   Circle "Circle_13" at 535,337 size 20x20
      Appearance <- "Data_Tank1_Heating_Cmd_ManCtrl"

screen "Mixing" 800x480
   TextField "Text field_26" at 286,251 size 194x23; Text 'Mixing phase control'
   TextField "Text field_27" at 182,285 size 83x23; Text 'Automat'
   TextField "Text field_28" at 182,303 size 70x23; Text 'Manual'
   TextField "Text field_29" at 343,294 size 51x23; Text 'Done'
   GraphicView "Graphic view_1" at 525,246 size 75x74; Picture "exit-png-cancel-cross-exit-remove-icon-512"
   Button "Button_26" at 520,248 size 76x81; TextOff 'Text'
      on Click: ActivateScreen("MainScr", 0)
   Button "Button_5" at 185,334 size 77x32; TextOff 'Aut'
      on Click: SetBit("Data_Tank1_Mixing_Cmd_AutCtrl")
   Button "Button_6" at 264,335 size 77x32; TextOff 'Man'
      on Click: SetBit("Data_Tank1_Mixing_Cmd_ManCtrl")
   Button "Button_12" at 186,371 size 77x32; TextOff 'Start'
      on Click: SetBit("Data_Tank1_Mixing_Cmd_StartMan")
   Button "Button_13" at 263,371 size 77x32; TextOff 'Stop'
      on Click: SetBit("Data_Tank1_Mixing_Cmd_StopMan")
   Button "Button_11" at 347,337 size 158x32; TextOff 'Reset Done'
      on Click: SetBit("Data_Tank1_Mixing_Cmd_ResetDone")
   Button "Button_14" at 350,371 size 77x32; TextOff 'Pause'
      on Click: SetBit("Data_Tank1_Mixing_Cmd_PauseMan")
   Button "Button_20" at 428,371 size 77x32; TextOff 'Rsume'
      on Click: SetBit("Data_Tank1_Mixing_Cmd_ResumeMan")
   Circle "Circle_5" at 445,291 size 35x35
      Appearance <- "Data_Tank1_Mixing_State_Done"
   Circle "Circle_6" at 290,285 size 20x20
      Appearance <- "Data_Tank1_Mixing_State_AutCtrl"
   Circle "Circle_7" at 290,309 size 20x20
      Appearance <- "Data_Tank1_Mixing_State_ManCtrl"
   SymbolLibrary "Symbol library_1" at 202,63 size 120x212
   SymbolLibrary "Symbol library_2" at 148,84 size 58x23
   SymbolLibrary "Symbol library_3" at 320,241 size 20x23
   Bar "Bar_1" at 204,63 size 117x211; MinimumValue 0; MaximumValue 2
      ProcessValue <- "Data_Tank1_WaterLevel_AIScaled"
   SymbolLibrary "Symbol library_4" at 55,31 size 94x80
      Appearance <- "Data_Tank1_ValveFill_State_StColor"
   IOField "I/O field_1" at 215,109 size 96x32; FormatPattern s9.99; Unit  m
      ProcessValue <- "Data_Tank1_WaterLevel_AIScaled"
   IOField "I/O field_2" at 216,143 size 96x32; FormatPattern 999.9; Unit  °C
      ProcessValue <- "Data_Tank1_WaterTemp_AIScaled"
   SymbolLibrary "Symbol library_6" at 226,190 size 71x61
      Appearance <- "Data_Tank1_Mixer_State_StateInt"
   Button "Button_1" at 7,233 size 77x32; TextOff 'Aut'
      on Click: SetBit("Data_Tank1_ValveFill_Cmd_AutCtrl")
   TextField "Text field_1" at 45,123 size 83x23; Text 'ValveFill'
   TextField "Text field_2" at 5,148 size 83x23; Text 'Automat'
   TextField "Text field_3" at 5,166 size 70x23; Text 'Manual'
   TextField "Text field_4" at 5,188 size 51x23; Text 'Open'
   TextField "Text field_5" at 5,206 size 65x23; Text 'Closed'
   Button "Button_2" at 86,233 size 77x32; TextOff 'Man'
      on Click: SetBit("Data_Tank1_ValveFill_Cmd_ManCtrl")
   Button "Button_3" at 7,267 size 77x32; TextOff 'Open'
      on Click: SetBit("Data_Tank1_ValveFill_Cmd_OpenMan")
   Button "Button_4" at 86,267 size 77x32; TextOff 'Close'
      on Click: SetBit("Data_Tank1_ValveFill_Cmd_CloseMan")
   TextField "Text field_6" at 450,99 size 104x23; Text 'ValveDrain'
   TextField "Text field_7" at 417,124 size 83x23; Text 'Automat'
   TextField "Text field_8" at 417,142 size 70x23; Text 'Manual'
   TextField "Text field_9" at 417,164 size 51x23; Text 'Open'
   TextField "Text field_10" at 417,182 size 65x23; Text 'Closed'
   Button "Button_9" at 187,378 size 77x32; TextOff 'Aut'
      on Click: SetBit("Data_Tank1_Mixer_Cmd_AutCtrl")
   TextField "Text field_11" at 234,284 size 56x23; Text 'Mixer'
   TextField "Text field_12" at 185,309 size 83x23; Text 'Automat'
   TextField "Text field_13" at 185,327 size 70x23; Text 'Manual'
   TextField "Text field_14" at 185,350 size 79x23; Text 'Running'
   Button "Button_10" at 266,378 size 77x32; TextOff 'Man'
      on Click: SetBit("Data_Tank1_Mixer_Cmd_ManCtrl")
   TextField "Text field_16" at 662,99 size 77x27; Text 'Phases'
   Button "Button_15" at 617,148 size 171x29; TextOff 'Menu filling'
      on Click: ActivateScreen("Filling", 0)
   TextField "Text field_17" at 668,124 size 61x23; Text 'Filling'
   SymbolicIOField "Symbolic I/O field_2" at 617,179 size 171x32; TextOn '1'; TextOff '0'; TextList "Phases"
      ProcessValue <- "Data_Tank1_Filling_State_Stateint"
   Button "Button_16" at 617,236 size 171x29; TextOff 'Menu draining'
      on Click: ActivateScreen("Draining", 0)
   TextField "Text field_18" at 660,213 size 82x23; Text 'Draining'
   SymbolicIOField "Symbolic I/O field_3" at 617,267 size 171x32; TextOn '1'; TextOff '0'; TextList "Phases"
      ProcessValue <- "Data_Tank1_Draining_State_StateInt"
   Button "Button_17" at 617,324 size 171x29; TextOff 'Menu mixing'
      on Click: ActivateScreen("Mixing", 0)
   TextField "Text field_19" at 669,301 size 65x23; Text 'Mixing'
   SymbolicIOField "Symbolic I/O field_4" at 617,355 size 171x32; TextOn '1'; TextOff '0'; TextList "Phases"
      ProcessValue <- "Data_Tank1_Mixing_State_StateInt"
   Button "Button_18" at 617,412 size 171x29; TextOff 'Menu heating'
      on Click: ActivateScreen("Heating", 0)
   TextField "Text field_20" at 665,390 size 76x23; Text 'Heating'
   SymbolicIOField "Symbolic I/O field_5" at 617,443 size 171x32; TextOn '1'; TextOff '0'; TextList "Phases"
      ProcessValue <- "Data_Tank1_Heating_State_StateInt"
   TextField "Text field_21" at 427,291 size 156x23; Text 'Heating element'
   TextField "Text field_22" at 418,316 size 83x23; Text 'Automat'
   TextField "Text field_23" at 418,334 size 70x23; Text 'Manual'
   TextField "Text field_24" at 422,356 size 157x23; Text 'Manual heat pwr'
   IOField "I/O field_3" at 447,377 size 96x32; FormatPattern 999.9; Unit  %
      ProcessValue <- "Data_Tank1_Heater_Param_HeatingPowerManual"
   TextField "Text field_25" at 422,408 size 160x23; Text 'Req temperature'
   Button "Button_27" at 335,12 size 130x66; TextOff 'Parameters tank 1'
      on Click: ActivateScreen("Parameters", 0)
   Circle "Circle_1" at 122,149 size 20x20
      Appearance <- "Data_Tank1_ValveFill_State_AutCtrl"
   Circle "Circle_2" at 122,169 size 20x20
      Appearance <- "Data_Tank1_ValveFill_State_ManCtrl"
   Circle "Circle_3" at 122,189 size 20x20
      Appearance <- "Data_Tank1_ValveFill_State_Open"
   Circle "Circle_4" at 122,209 size 20x20
      Appearance <- "Data_Tank1_ValveFill_State_Closed"
   Circle "Circle_9" at 302,310 size 20x20
      Appearance <- "Data_Tank1_Mixer_State_AutCtrl"
   Circle "Circle_10" at 302,330 size 20x20
      Appearance <- "Data_Tank1_Mixer_State_ManCtrl"
   Circle "Circle_12" at 302,354 size 20x20
      Appearance <- "Data_Tank1_Mixer_State_Run"
   Circle "Circle_11" at 535,317 size 20x20
      Appearance <- "Data_Tank1_Heating_Cmd_AutCtrl"
   Circle "Circle_13" at 535,337 size 20x20
      Appearance <- "Data_Tank1_Heating_Cmd_ManCtrl"
   TextField "Text field_30" at 427,285 size 156x23; Text 'Heating element'
   TextField "Text field_31" at 418,310 size 83x23; Text 'Automat'
   TextField "Text field_32" at 418,328 size 70x23; Text 'Manual'
   TextField "Text field_33" at 422,350 size 157x23; Text 'Manual heat pwr'
   Circle "Circle_17" at 535,311 size 20x20
      Appearance <- "Data_Tank1_Heater_State_AutCtrl"
   Circle "Circle_18" at 535,331 size 20x20
      Appearance <- "Data_Tank1_Heater_State_ManCtrl"
   IOField "I/O field_4" at 447,371 size 96x32; FormatPattern 999.9; Unit  %
      ProcessValue <- "Data_Tank1_Heater_Param_HeatingPowerManual"

